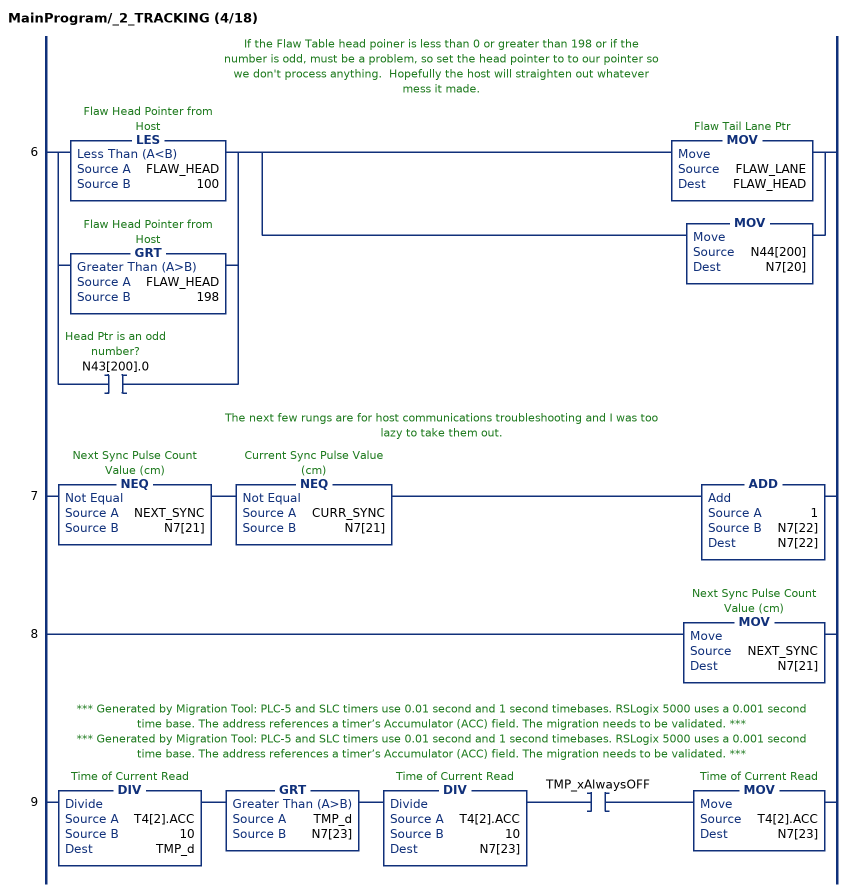
   // If the Flaw Table head poiner is less than 0 or greater than 198 or if the
   // number is odd, must be a problem, so set the head pointer to to our pointer so
   // we don't process anything.  Hopefully the host will straighten out whatever
   // mess it made.
   6: [LES(FLAW_HEAD,100) ,GRT(FLAW_HEAD,198) ,XIC(N43[200].0) ][MOV(FLAW_LANE,FLAW_HEAD) ,MOV(N44[200],N7[20]) ];
   // The next few rungs are for host communications troubleshooting and I was too
   // lazy to take them out.
   7: NEQ(NEXT_SYNC,N7[21])NEQ(CURR_SYNC,N7[21])ADD(1,N7[22],N7[22]);
   8: MOV(NEXT_SYNC,N7[21]);
   // *** Generated by Migration Tool: PLC-5 and SLC timers use 0.01 second and 1 second timebases. RSLogix 5000 uses a 0.001 second time base. The address references a timer’s Accumulator (ACC) field. The migration needs to be validated. ***
   // *** Generated by Migration Tool: PLC-5 and SLC timers use 0.01 second and 1 second timebases. RSLogix 5000 uses a 0.001 second time base. The address references a timer’s Accumulator (ACC) field. The migration needs to be validated. ***
   9: DIV(T4[2].ACC,10,TMP_d)GRT(TMP_d,N7[23])DIV(T4[2].ACC,10,N7[23])XIC(TMP_xAlwaysOFF)MOV(T4[2].ACC,N7[23]);
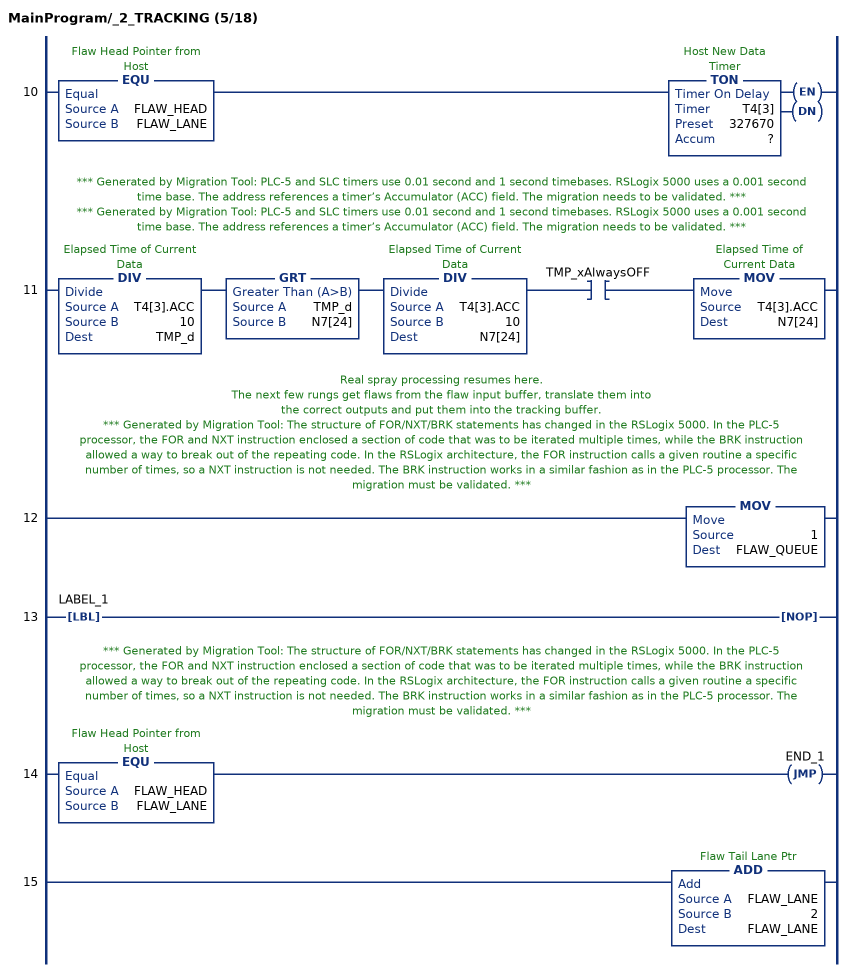
   10: EQU(FLAW_HEAD,FLAW_LANE)TON(T4[3],?,?);
   // *** Generated by Migration Tool: PLC-5 and SLC timers use 0.01 second and 1 second timebases. RSLogix 5000 uses a 0.001 second time base. The address references a timer’s Accumulator (ACC) field. The migration needs to be validated. ***
   // *** Generated by Migration Tool: PLC-5 and SLC timers use 0.01 second and 1 second timebases. RSLogix 5000 uses a 0.001 second time base. The address references a timer’s Accumulator (ACC) field. The migration needs to be validated. ***
   11: DIV(T4[3].ACC,10,TMP_d)GRT(TMP_d,N7[24])DIV(T4[3].ACC,10,N7[24])XIC(TMP_xAlwaysOFF)MOV(T4[3].ACC,N7[24]);
   // Real spray processing resumes here.
   // The next few rungs get flaws from the flaw input buffer, translate them into
   // the correct outputs and put them into the tracking buffer.
   // *** Generated by Migration Tool: The structure of FOR/NXT/BRK statements has changed in the RSLogix 5000. In the PLC-5 processor, the FOR and NXT instruction enclosed a section of code that was to be iterated multiple times, while the BRK instruction allowed a way to break out of the repeating code. In the RSLogix architecture, the FOR instruction calls a given routine a specific number of times, so a NXT instruction is not needed. The BRK instruction works in a similar fashion as in the PLC-5 processor. The migration must be validated. ***
   12: MOV(1,FLAW_QUEUE);
   13: LBL(LABEL_1)NOP();
   // *** Generated by Migration Tool: The structure of FOR/NXT/BRK statements has changed in the RSLogix 5000. In the PLC-5 processor, the FOR and NXT instruction enclosed a section of code that was to be iterated multiple times, while the BRK instruction allowed a way to break out of the repeating code. In the RSLogix architecture, the FOR instruction calls a given routine a specific number of times, so a NXT instruction is not needed. The BRK instruction works in a similar fashion as in the PLC-5 processor. The migration must be validated. ***
   14: EQU(FLAW_HEAD,FLAW_LANE)JMP(END_1);
   15: ADD(FLAW_LANE,2,FLAW_LANE);
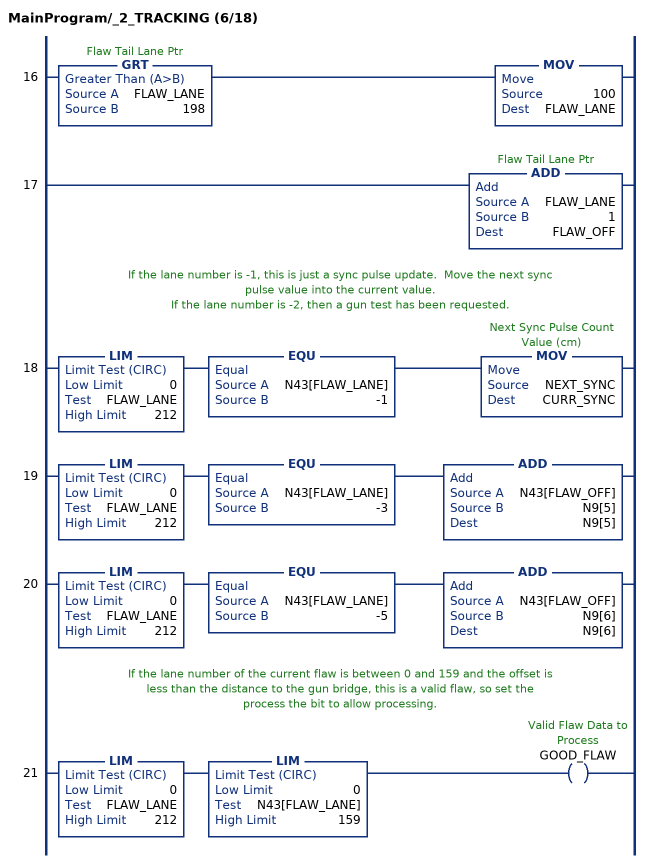
   16: GRT(FLAW_LANE,198)MOV(100,FLAW_LANE);
   17: ADD(FLAW_LANE,1,FLAW_OFF);
   // If the lane number is -1, this is just a sync pulse update.  Move the next sync
   // pulse value into the current value.
   // If the lane number is -2, then a gun test has been requested.
   18: LIM(0,FLAW_LANE,212)EQU(N43[FLAW_LANE],-1)MOV(NEXT_SYNC,CURR_SYNC);
   19: LIM(0,FLAW_LANE,212)EQU(N43[FLAW_LANE],-3)ADD(N43[FLAW_OFF],N9[5],N9[5]);
   20: LIM(0,FLAW_LANE,212)EQU(N43[FLAW_LANE],-5)ADD(N43[FLAW_OFF],N9[6],N9[6]);
   // If the lane number of the current flaw is between 0 and 159 and the offset is
   // less than the distance to the gun bridge, this is a valid flaw, so set the
   // process the bit to allow processing.
   21: LIM(0,FLAW_LANE,212)LIM(0,N43[FLAW_LANE],159)OTE(GOOD_FLAW);
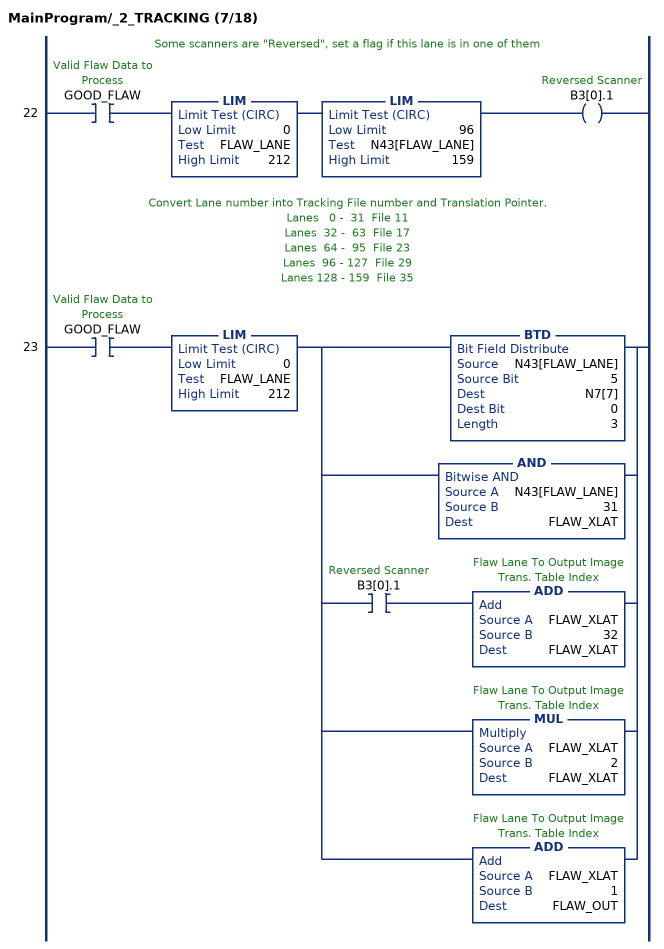
   // Some scanners are "Reversed", set a flag if this lane is in one of them
   22: XIC(GOOD_FLAW)LIM(0,FLAW_LANE,212)LIM(96,N43[FLAW_LANE],159)OTE(B3[0].1);
   // Convert Lane number into Tracking File number and Translation Pointer.
   //      Lanes   0 -  31  File 11
   //      Lanes  32 -  63  File 17
   //      Lanes  64 -  95  File 23
   //      Lanes  96 - 127  File 29
   //      Lanes 128 - 159  File 35
   23: XIC(GOOD_FLAW)LIM(0,FLAW_LANE,212)[BTD(N43[FLAW_LANE],5,N7[7],0,3) ,AND(N43[FLAW_LANE],31,FLAW_XLAT) ,XIC(B3[0].1) ADD(FLAW_XLAT,32,FLAW_XLAT) ,MUL(FLAW_XLAT,2,FLAW_XLAT) ,ADD(FLAW_XLAT,1,FLAW_OUT) ];
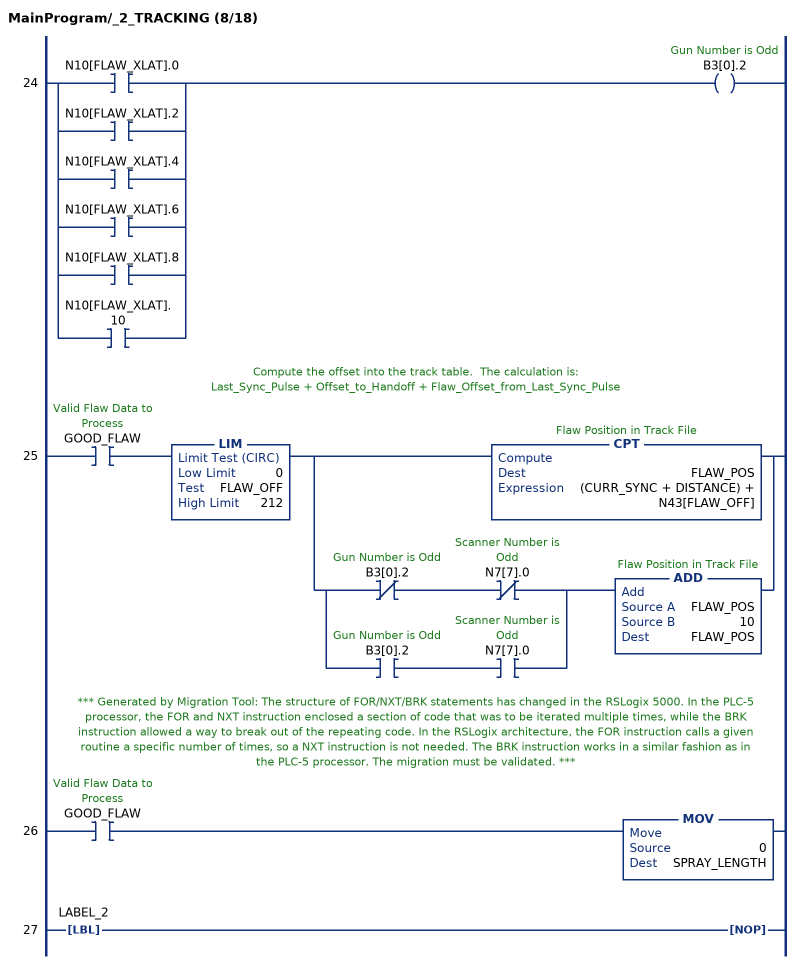
   24: [XIC(N10[FLAW_XLAT].0) ,XIC(N10[FLAW_XLAT].2) ,XIC(N10[FLAW_XLAT].4) ,XIC(N10[FLAW_XLAT].6) ,XIC(N10[FLAW_XLAT].8) ,XIC(N10[FLAW_XLAT].10) ]OTE(B3[0].2);
   // Compute the offset into the track table.  The calculation is:
   //    Last_Sync_Pulse + Offset_to_Handoff + Flaw_Offset_from_Last_Sync_Pulse
   25: XIC(GOOD_FLAW)LIM(0,FLAW_OFF,212)[CPT(FLAW_POS,(CURR_SYNC + DISTANCE) + N43[FLAW_OFF]) ,[XIO(B3[0].2) XIO(N7[7].0) ,XIC(B3[0].2) XIC(N7[7].0) ] ADD(FLAW_POS,10,FLAW_POS) ];
   // *** Generated by Migration Tool: The structure of FOR/NXT/BRK statements has changed in the RSLogix 5000. In the PLC-5 processor, the FOR and NXT instruction enclosed a section of code that was to be iterated multiple times, while the BRK instruction allowed a way to break out of the repeating code. In the RSLogix architecture, the FOR instruction calls a given routine a specific number of times, so a NXT instruction is not needed. The BRK instruction works in a similar fashion as in the PLC-5 processor. The migration must be validated. ***
   26: XIC(GOOD_FLAW)MOV(0,SPRAY_LENGTH);
   27: LBL(LABEL_2)NOP();
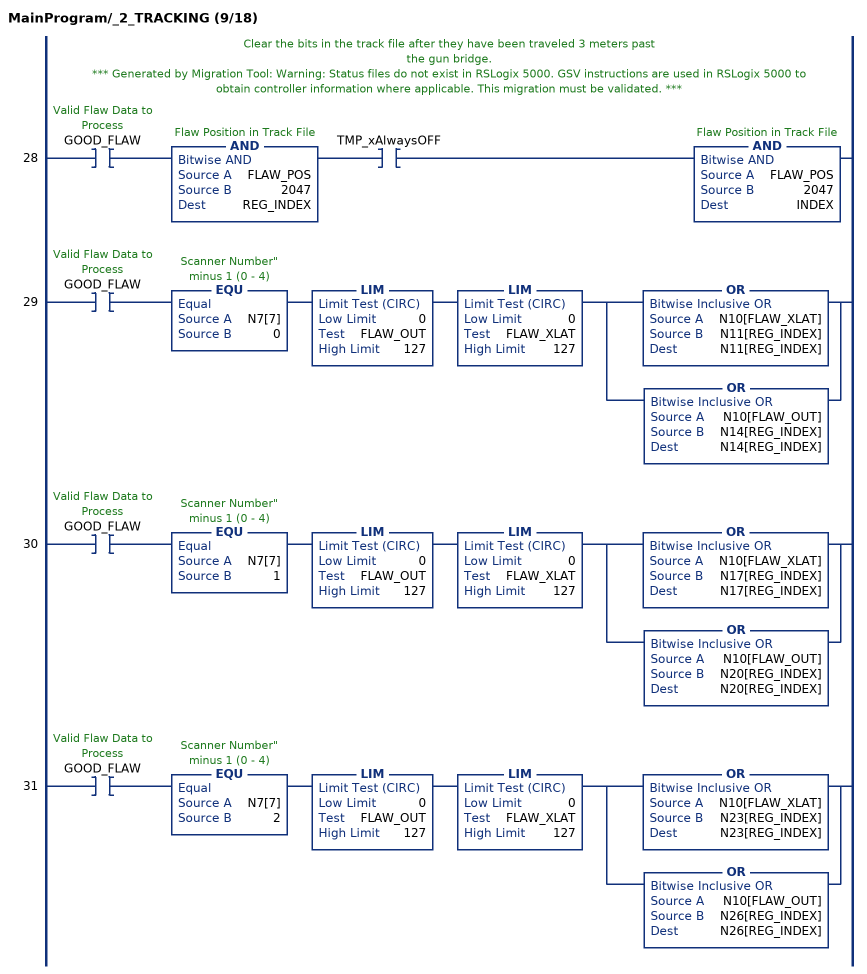
   // Clear the bits in the track file after they have been traveled 3 meters past
   // the gun bridge.
   // *** Generated by Migration Tool: Warning: Status files do not exist in RSLogix 5000. GSV instructions are used in RSLogix 5000 to obtain controller information where applicable. This migration must be validated. ***
   28: XIC(GOOD_FLAW)AND(FLAW_POS,2047,REG_INDEX)XIC(TMP_xAlwaysOFF)AND(FLAW_POS,2047,INDEX);
   29: XIC(GOOD_FLAW)EQU(N7[7],0)LIM(0,FLAW_OUT,127)LIM(0,FLAW_XLAT,127)[OR(N10[FLAW_XLAT],N11[REG_INDEX],N11[REG_INDEX]) ,OR(N10[FLAW_OUT],N14[REG_INDEX],N14[REG_INDEX]) ];
   30: XIC(GOOD_FLAW)EQU(N7[7],1)LIM(0,FLAW_OUT,127)LIM(0,FLAW_XLAT,127)[OR(N10[FLAW_XLAT],N17[REG_INDEX],N17[REG_INDEX]) ,OR(N10[FLAW_OUT],N20[REG_INDEX],N20[REG_INDEX]) ];
   31: XIC(GOOD_FLAW)EQU(N7[7],2)LIM(0,FLAW_OUT,127)LIM(0,FLAW_XLAT,127)[OR(N10[FLAW_XLAT],N23[REG_INDEX],N23[REG_INDEX]) ,OR(N10[FLAW_OUT],N26[REG_INDEX],N26[REG_INDEX]) ];
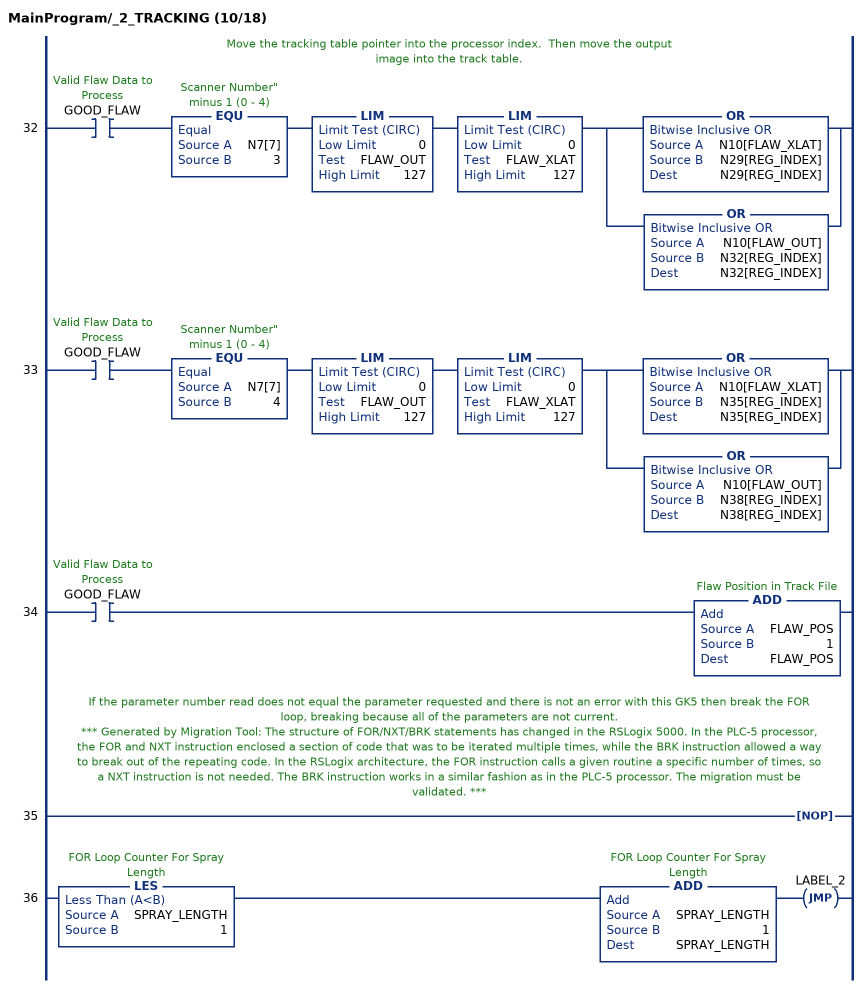
   // Move the tracking table pointer into the processor index.  Then move the output
   // image into the track table.
   32: XIC(GOOD_FLAW)EQU(N7[7],3)LIM(0,FLAW_OUT,127)LIM(0,FLAW_XLAT,127)[OR(N10[FLAW_XLAT],N29[REG_INDEX],N29[REG_INDEX]) ,OR(N10[FLAW_OUT],N32[REG_INDEX],N32[REG_INDEX]) ];
   33: XIC(GOOD_FLAW)EQU(N7[7],4)LIM(0,FLAW_OUT,127)LIM(0,FLAW_XLAT,127)[OR(N10[FLAW_XLAT],N35[REG_INDEX],N35[REG_INDEX]) ,OR(N10[FLAW_OUT],N38[REG_INDEX],N38[REG_INDEX]) ];
   34: XIC(GOOD_FLAW)ADD(FLAW_POS,1,FLAW_POS);
   // If the parameter number read does not equal the parameter requested and there is not an error with this GK5 then break the FOR
   // loop, breaking because all of the parameters are not current.
   // *** Generated by Migration Tool: The structure of FOR/NXT/BRK statements has changed in the RSLogix 5000. In the PLC-5 processor, the FOR and NXT instruction enclosed a section of code that was to be iterated multiple times, while the BRK instruction allowed a way to break out of the repeating code. In the RSLogix architecture, the FOR instruction calls a given routine a specific number of times, so a NXT instruction is not needed. The BRK instruction works in a similar fashion as in the PLC-5 processor. The migration must be validated. ***
   35: NOP();
   36: LES(SPRAY_LENGTH,1)ADD(SPRAY_LENGTH,1,SPRAY_LENGTH)JMP(LABEL_2);
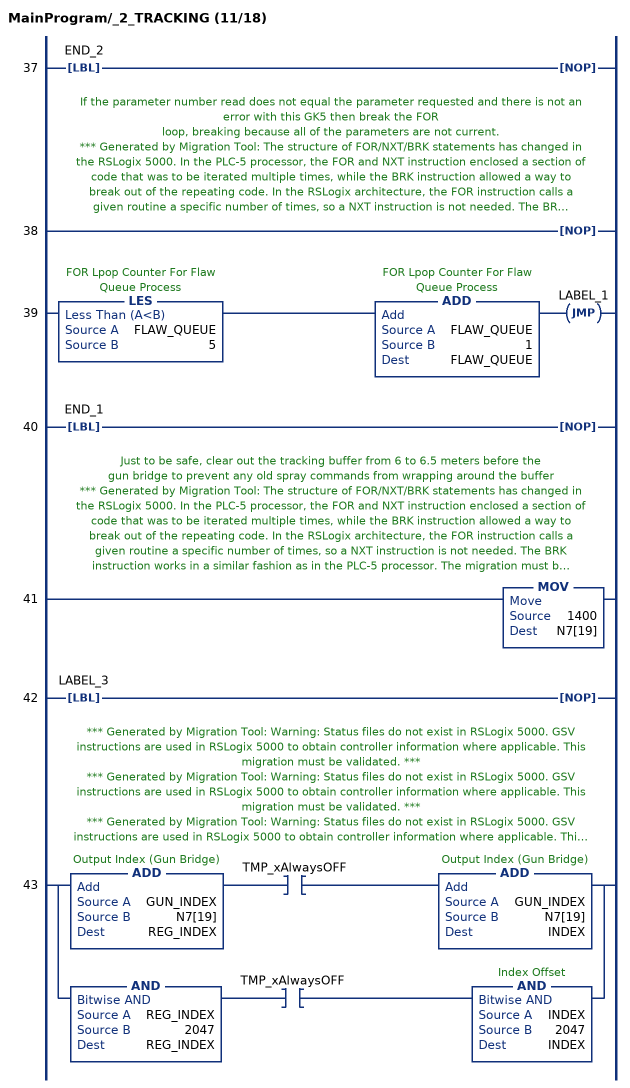
   37: LBL(END_2)NOP();
   // If the parameter number read does not equal the parameter requested and there is not an error with this GK5 then break the FOR
   // loop, breaking because all of the parameters are not current.
   // *** Generated by Migration Tool: The structure of FOR/NXT/BRK statements has changed in the RSLogix 5000. In the PLC-5 processor, the FOR and NXT instruction enclosed a section of code that was to be iterated multiple times, while the BRK instruction allowed a way to break out of the repeating code. In the RSLogix architecture, the FOR instruction calls a given routine a specific number of times, so a NXT instruction is not needed. The BRK instruction works in a similar fashion as in the PLC-5 processor. The migration must be validated. ***
   38: NOP();
   39: LES(FLAW_QUEUE,5)ADD(FLAW_QUEUE,1,FLAW_QUEUE)JMP(LABEL_1);
   40: LBL(END_1)NOP();
   // Just to be safe, clear out the tracking buffer from 6 to 6.5 meters before the
   // gun bridge to prevent any old spray commands from wrapping around the buffer
   // *** Generated by Migration Tool: The structure of FOR/NXT/BRK statements has changed in the RSLogix 5000. In the PLC-5 processor, the FOR and NXT instruction enclosed a section of code that was to be iterated multiple times, while the BRK instruction allowed a way to break out of the repeating code. In the RSLogix architecture, the FOR instruction calls a given routine a specific number of times, so a NXT instruction is not needed. The BRK instruction works in a similar fashion as in the PLC-5 processor. The migration must be validated. ***
   41: MOV(1400,N7[19]);
   42: LBL(LABEL_3)NOP();
   // *** Generated by Migration Tool: Warning: Status files do not exist in RSLogix 5000. GSV instructions are used in RSLogix 5000 to obtain controller information where applicable. This migration must be validated. ***
   // *** Generated by Migration Tool: Warning: Status files do not exist in RSLogix 5000. GSV instructions are used in RSLogix 5000 to obtain controller information where applicable. This migration must be validated. ***
   // *** Generated by Migration Tool: Warning: Status files do not exist in RSLogix 5000. GSV instructions are used in RSLogix 5000 to obtain controller information where applicable. This migration must be validated. ***
   43: [ADD(GUN_INDEX,N7[19],REG_INDEX) XIC(TMP_xAlwaysOFF) ADD(GUN_INDEX,N7[19],INDEX) ,AND(REG_INDEX,2047,REG_INDEX) XIC(TMP_xAlwaysOFF) AND(INDEX,2047,INDEX) ];
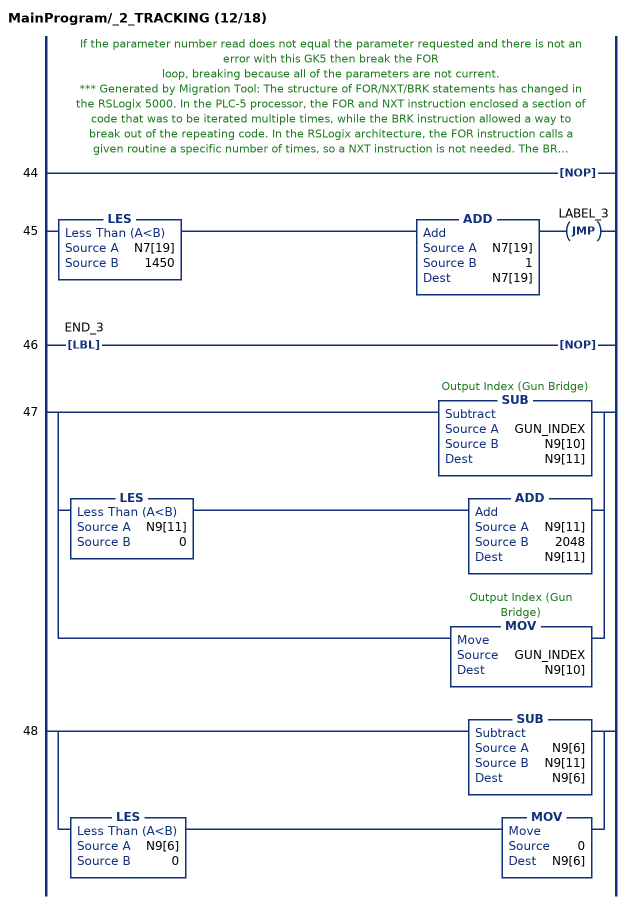
   // If the parameter number read does not equal the parameter requested and there is not an error with this GK5 then break the FOR
   // loop, breaking because all of the parameters are not current.
   // *** Generated by Migration Tool: The structure of FOR/NXT/BRK statements has changed in the RSLogix 5000. In the PLC-5 processor, the FOR and NXT instruction enclosed a section of code that was to be iterated multiple times, while the BRK instruction allowed a way to break out of the repeating code. In the RSLogix architecture, the FOR instruction calls a given routine a specific number of times, so a NXT instruction is not needed. The BRK instruction works in a similar fashion as in the PLC-5 processor. The migration must be validated. ***
   44: NOP();
   45: LES(N7[19],1450)ADD(N7[19],1,N7[19])JMP(LABEL_3);
   46: LBL(END_3)NOP();
   47: [SUB(GUN_INDEX,N9[10],N9[11]) ,LES(N9[11],0) ADD(N9[11],2048,N9[11]) ,MOV(GUN_INDEX,N9[10]) ];
   48: [SUB(N9[6],N9[11],N9[6]) ,LES(N9[6],0) MOV(0,N9[6]) ];
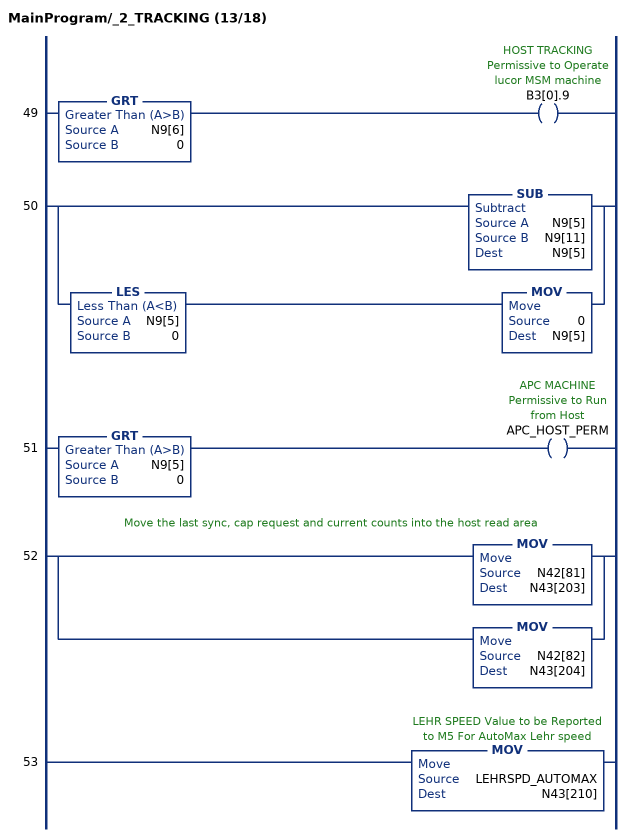
   49: GRT(N9[6],0)OTE(B3[0].9);
   50: [SUB(N9[5],N9[11],N9[5]) ,LES(N9[5],0) MOV(0,N9[5]) ];
   51: GRT(N9[5],0)OTE(APC_HOST_PERM);
   // Move the last sync, cap request and current counts into the host read area
   52: [MOV(N42[81],N43[203]) ,MOV(N42[82],N43[204]) ];
   53: MOV(LEHRSPD_AUTOMAX,N43[210]);
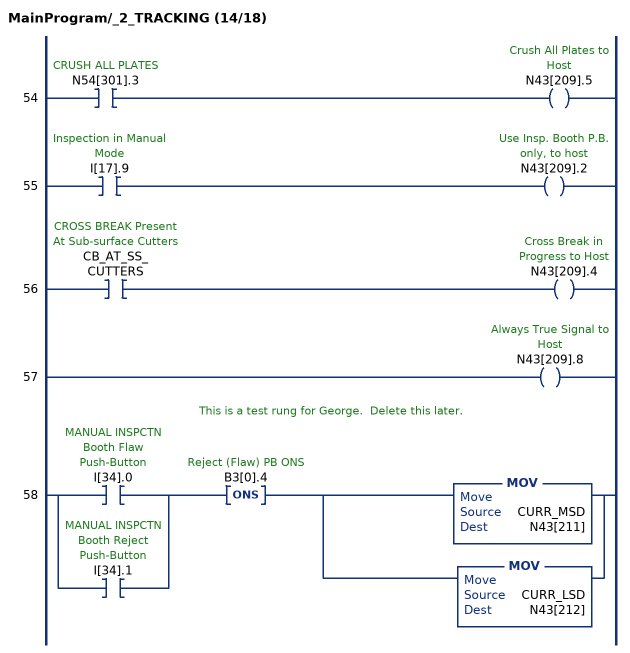
   54: XIC(N54[301].3)OTE(N43[209].5);
   55: XIC(I[17].9)OTE(N43[209].2);
   56: XIC(CB_AT_SS_CUTTERS)OTE(N43[209].4);
   57: OTE(N43[209].8);
   // This is a test rung for George.  Delete this later.
   58: [XIC(I[34].0) ,XIC(I[34].1) ]ONS(B3[0].4)[MOV(CURR_MSD,N43[211]) ,MOV(CURR_LSD,N43[212]) ];
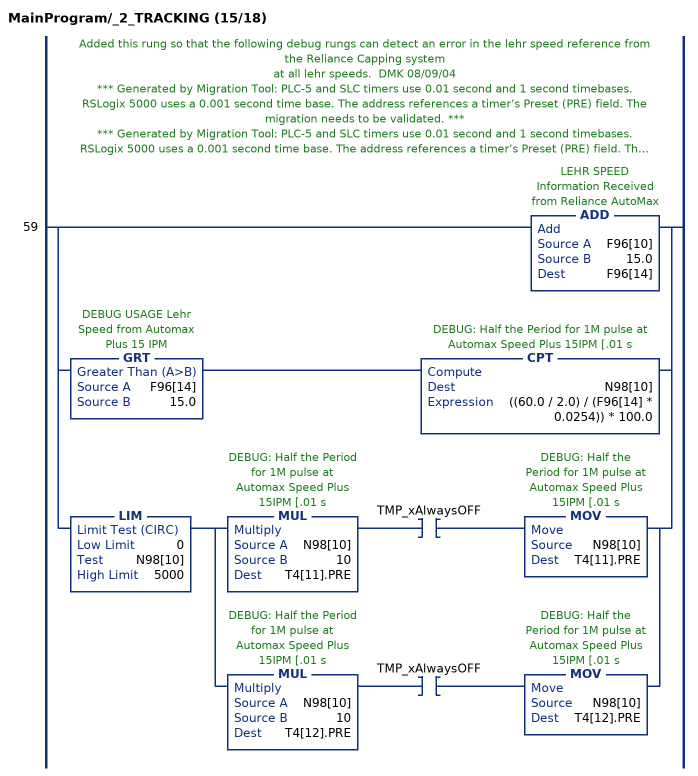
   // Added this rung so that the following debug rungs can detect an error in the lehr speed reference from the Reliance Capping system
   // at all lehr speeds.  DMK 08/09/04
   // *** Generated by Migration Tool: PLC-5 and SLC timers use 0.01 second and 1 second timebases. RSLogix 5000 uses a 0.001 second time base. The address references a timer’s Preset (PRE) field. The migration needs to be validated. ***
   // *** Generated by Migration Tool: PLC-5 and SLC timers use 0.01 second and 1 second timebases. RSLogix 5000 uses a 0.001 second time base. The address references a timer’s Preset (PRE) field. The migration needs to be validated. ***
   59: [ADD(F96[10],15.0,F96[14]) ,GRT(F96[14],15.0) CPT(N98[10],((60.0 / 2.0) / (F96[14] * 0.0254)) * 100.0) ,LIM(0,N98[10],5000) [MUL(N98[10],10,T4[11].PRE) XIC(TMP_xAlwaysOFF) MOV(N98[10],T4[11].PRE) ,MUL(N98[10],10,T4[12].PRE) XIC(TMP_xAlwaysOFF) MOV(N98[10],T4[12].PRE) ] ];
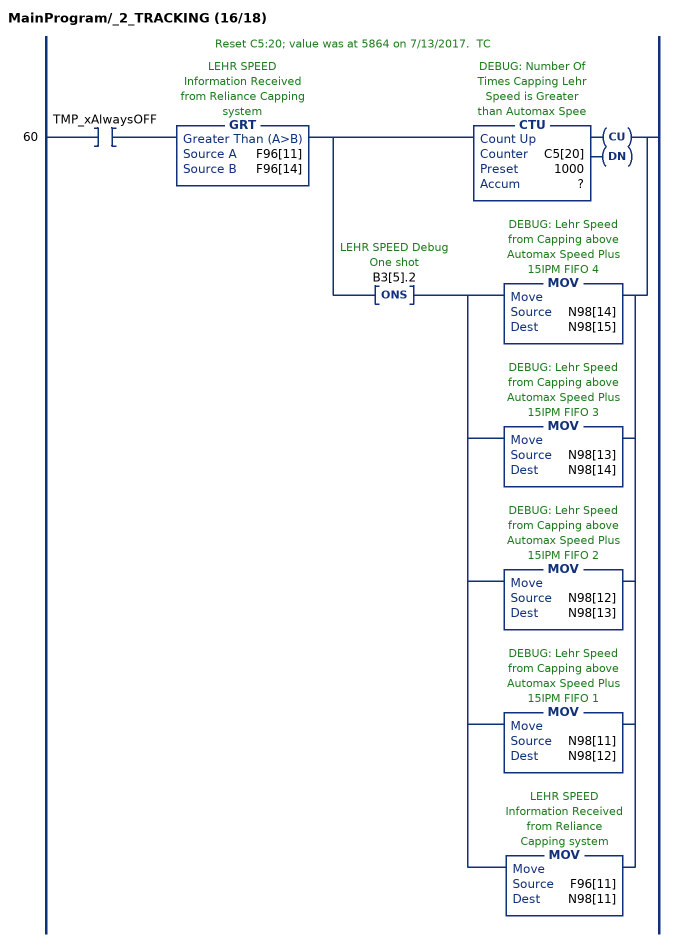
   // Reset C5:20; value was at 5864 on 7/13/2017.  TC
   60: XIC(TMP_xAlwaysOFF)GRT(F96[11],F96[14])[CTU(C5[20],?,?) ,ONS(B3[5].2) [MOV(N98[14],N98[15]) ,MOV(N98[13],N98[14]) ,MOV(N98[12],N98[13]) ,MOV(N98[11],N98[12]) ,MOV(F96[11],N98[11]) ] ];
